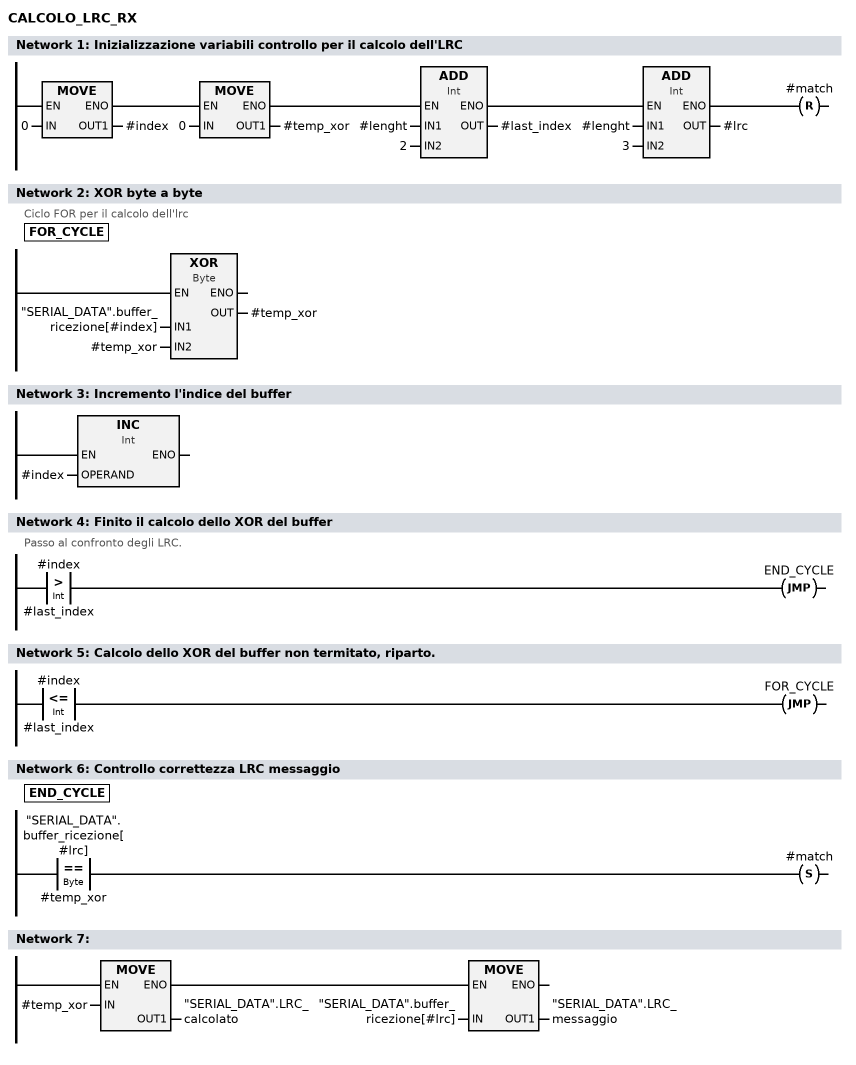
   RUNG wire#powerrail
      Move(in := 0, out1 => #index)
      Move(in := 0, out1 => #temp_xor)
      { S7_Templates := "SrcType := Int" } Add(in1 := #lenght, in2 := 2, out => #last_index)
      { S7_Templates := "SrcType := Int" } Add(in1 := #lenght, in2 := 3, out => #lrc)
      R_Coil( #match )
   END_RUNG
   // the same network as SCL:
   #index := 0;
   #temp_xor := 0;
   #last_index := #lenght + 2;
   #lrc := #lenght + 3;
   #match := FALSE;
END_REGION

REGION Network 2: XOR byte a byte
   // Ciclo FOR per il calcolo dell'lrc
   // no checked SCL form for this network; see the picture
END_REGION

REGION Network 3: Incremento l'indice del buffer
   RUNG wire#powerrail
      { S7_Templates := "DestType := Int" } Inc( #index )
   END_RUNG
   // the same network as SCL:
   #index := #index + 1;
END_REGION

REGION Network 4: Finito il calcolo dello XOR del buffer
   // Passo al confronto degli LRC.
   RUNG wire#powerrail
      { S7_Templates := "SrcType := Int" } GT_Contact(in1 := #index, in2 := #last_index)
      JumpCoil( END_CYCLE )
   END_RUNG
   // the same network as SCL:
   IF #index > #last_index THEN GOTO END_CYCLE; END_IF;
END_REGION

REGION Network 5: Calcolo dello XOR del buffer non termitato, riparto.
   RUNG wire#powerrail
      { S7_Templates := "SrcType := Int" } LE_Contact(in1 := #index, in2 := #last_index)
      JumpCoil( FOR_CYCLE )
   END_RUNG
   // the same network as SCL:
   IF #index <= #last_index THEN GOTO FOR_CYCLE; END_IF;
END_REGION

REGION Network 6: Controllo correttezza LRC messaggio
   Label( END_CYCLE )
   RUNG wire#powerrail
      { S7_Templates := "SrcType := Byte" } EQ_Contact(in1 := "SERIAL_DATA".buffer_ricezione[#lrc], in2 := #temp_xor)
      S_Coil( #match )
   END_RUNG
   // the same network as SCL:
   END_CYCLE:
   IF "SERIAL_DATA".buffer_ricezione[#lrc] = #temp_xor THEN #match := TRUE; END_IF;
END_REGION

REGION Network 7
   RUNG wire#powerrail
      Move(in := #temp_xor, out1 => "SERIAL_DATA".LRC_calcolato)
      Move(in := "SERIAL_DATA".buffer_ricezione[#lrc], out1 => "SERIAL_DATA".LRC_messaggio)
   END_RUNG
   // the same network as SCL:
   "SERIAL_DATA".LRC_calcolato := #temp_xor;
   "SERIAL_DATA".LRC_messaggio := "SERIAL_DATA".buffer_ricezione[#lrc];
END_REGION
END_FUNCTION

FUNCTION "RESET_ALLARMI" : Void   // FC7, LAD
TITLE = RESET ALLARMI
{ S7_Optimized_Access := 'FALSE' }
VERSION : 0.1
BEGIN

REGION Network 1: Azzero i contatori di fault Amplificatori
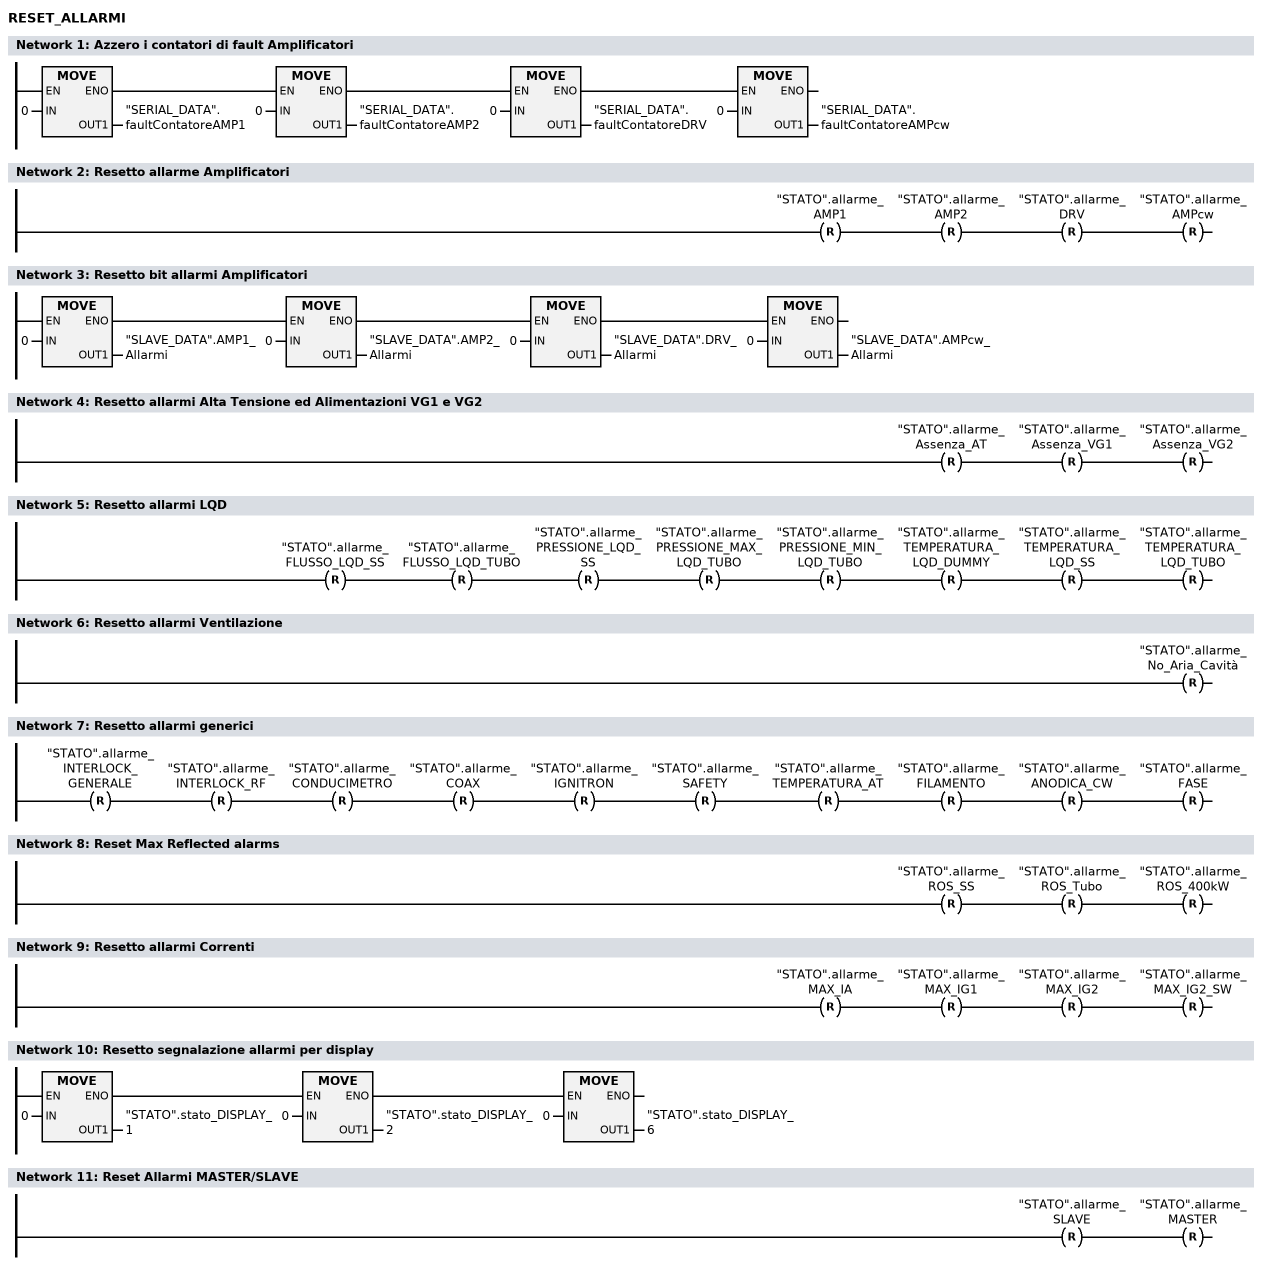
   RUNG wire#powerrail
      Move(in := 0, out1 => "SERIAL_DATA".faultContatoreAMP1)
      Move(in := 0, out1 => "SERIAL_DATA".faultContatoreAMP2)
      Move(in := 0, out1 => "SERIAL_DATA".faultContatoreDRV)
      Move(in := 0, out1 => "SERIAL_DATA".faultContatoreAMPcw)
   END_RUNG
   // the same network as SCL:
   "SERIAL_DATA".faultContatoreAMP1 := 0;
   "SERIAL_DATA".faultContatoreAMP2 := 0;
   "SERIAL_DATA".faultContatoreDRV := 0;
   "SERIAL_DATA".faultContatoreAMPcw := 0;
END_REGION

REGION Network 2: Resetto allarme Amplificatori
   RUNG wire#powerrail
      R_Coil( "STATO".allarme_AMP1 )
      R_Coil( "STATO".allarme_AMP2 )
      R_Coil( "STATO".allarme_DRV )
      R_Coil( "STATO".allarme_AMPcw )
   END_RUNG
   // the same network as SCL:
   "STATO".allarme_AMP1 := FALSE;
   "STATO".allarme_AMP2 := FALSE;
   "STATO".allarme_DRV := FALSE;
   "STATO".allarme_AMPcw := FALSE;
END_REGION

REGION Network 3: Resetto bit allarmi Amplificatori
   RUNG wire#powerrail
      Move(in := 0, out1 => "SLAVE_DATA".AMP1_Allarmi)
      Move(in := 0, out1 => "SLAVE_DATA".AMP2_Allarmi)
      Move(in := 0, out1 => "SLAVE_DATA".DRV_Allarmi)
      Move(in := 0, out1 => "SLAVE_DATA".AMPcw_Allarmi)
   END_RUNG
   // the same network as SCL:
   "SLAVE_DATA".AMP1_Allarmi := 0;
   "SLAVE_DATA".AMP2_Allarmi := 0;
   "SLAVE_DATA".DRV_Allarmi := 0;
   "SLAVE_DATA".AMPcw_Allarmi := 0;
END_REGION

REGION Network 4: Resetto allarmi Alta Tensione ed Alimentazioni VG1 e VG2
   RUNG wire#powerrail
      R_Coil( "STATO".allarme_Assenza_AT )
      R_Coil( "STATO".allarme_Assenza_VG1 )
      R_Coil( "STATO".allarme_Assenza_VG2 )
   END_RUNG
   // the same network as SCL:
   "STATO".allarme_Assenza_AT := FALSE;
   "STATO".allarme_Assenza_VG1 := FALSE;
   "STATO".allarme_Assenza_VG2 := FALSE;
END_REGION

REGION Network 5: Resetto allarmi LQD
   RUNG wire#powerrail
      R_Coil( "STATO".allarme_FLUSSO_LQD_SS )
      R_Coil( "STATO".allarme_FLUSSO_LQD_TUBO )
      R_Coil( "STATO".allarme_PRESSIONE_LQD_SS )
      R_Coil( "STATO".allarme_PRESSIONE_MAX_LQD_TUBO )
      R_Coil( "STATO".allarme_PRESSIONE_MIN_LQD_TUBO )
      R_Coil( "STATO".allarme_TEMPERATURA_LQD_DUMMY )
      R_Coil( "STATO".allarme_TEMPERATURA_LQD_SS )
      R_Coil( "STATO".allarme_TEMPERATURA_LQD_TUBO )
   END_RUNG
   // the same network as SCL:
   "STATO".allarme_FLUSSO_LQD_SS := FALSE;
   "STATO".allarme_FLUSSO_LQD_TUBO := FALSE;
   "STATO".allarme_PRESSIONE_LQD_SS := FALSE;
   "STATO".allarme_PRESSIONE_MAX_LQD_TUBO := FALSE;
   "STATO".allarme_PRESSIONE_MIN_LQD_TUBO := FALSE;
   "STATO".allarme_TEMPERATURA_LQD_DUMMY := FALSE;
   "STATO".allarme_TEMPERATURA_LQD_SS := FALSE;
   "STATO".allarme_TEMPERATURA_LQD_TUBO := FALSE;
END_REGION

REGION Network 6: Resetto allarmi Ventilazione
   RUNG wire#powerrail
      R_Coil( "STATO".allarme_No_Aria_Cavità )
   END_RUNG
   // the same network as SCL:
   "STATO".allarme_No_Aria_Cavità := FALSE;
END_REGION

REGION Network 7: Resetto allarmi generici
   RUNG wire#powerrail
      R_Coil( "STATO".allarme_INTERLOCK_GENERALE )
      R_Coil( "STATO".allarme_INTERLOCK_RF )
      R_Coil( "STATO".allarme_CONDUCIMETRO )
      R_Coil( "STATO".allarme_COAX )
      R_Coil( "STATO".allarme_IGNITRON )
      R_Coil( "STATO".allarme_SAFETY )
      R_Coil( "STATO".allarme_TEMPERATURA_AT )
      R_Coil( "STATO".allarme_FILAMENTO )
      R_Coil( "STATO".allarme_ANODICA_CW )
      R_Coil( "STATO".allarme_FASE )
   END_RUNG
   // the same network as SCL:
   "STATO".allarme_INTERLOCK_GENERALE := FALSE;
   "STATO".allarme_INTERLOCK_RF := FALSE;
   "STATO".allarme_CONDUCIMETRO := FALSE;
   "STATO".allarme_COAX := FALSE;
   "STATO".allarme_IGNITRON := FALSE;
   "STATO".allarme_SAFETY := FALSE;
   "STATO".allarme_TEMPERATURA_AT := FALSE;
   "STATO".allarme_FILAMENTO := FALSE;
   "STATO".allarme_ANODICA_CW := FALSE;
   "STATO".allarme_FASE := FALSE;
END_REGION

REGION Network 8: Reset Max Reflected alarms
   RUNG wire#powerrail
      R_Coil( "STATO".allarme_ROS_SS )
      R_Coil( "STATO".allarme_ROS_Tubo )
      R_Coil( "STATO".allarme_ROS_400kW )
   END_RUNG
   // the same network as SCL:
   "STATO".allarme_ROS_SS := FALSE;
   "STATO".allarme_ROS_Tubo := FALSE;
   "STATO".allarme_ROS_400kW := FALSE;
END_REGION

REGION Network 9: Resetto allarmi Correnti
   RUNG wire#powerrail
      R_Coil( "STATO".allarme_MAX_IA )
      R_Coil( "STATO".allarme_MAX_IG1 )
      R_Coil( "STATO".allarme_MAX_IG2 )
      R_Coil( "STATO".allarme_MAX_IG2_SW )
   END_RUNG
   // the same network as SCL:
   "STATO".allarme_MAX_IA := FALSE;
   "STATO".allarme_MAX_IG1 := FALSE;
   "STATO".allarme_MAX_IG2 := FALSE;
   "STATO".allarme_MAX_IG2_SW := FALSE;
END_REGION

REGION Network 10: Resetto segnalazione allarmi per display
   RUNG wire#powerrail
      Move(in := 0, out1 => "STATO".stato_DISPLAY_1)
      Move(in := 0, out1 => "STATO".stato_DISPLAY_2)
      Move(in := 0, out1 => "STATO".stato_DISPLAY_6)
   END_RUNG
   // the same network as SCL:
   "STATO".stato_DISPLAY_1 := 0;
   "STATO".stato_DISPLAY_2 := 0;
   "STATO".stato_DISPLAY_6 := 0;
END_REGION

REGION Network 11: Reset Allarmi MASTER/SLAVE
   RUNG wire#powerrail
      R_Coil( "STATO".allarme_SLAVE )
      R_Coil( "STATO".allarme_MASTER )
   END_RUNG
   // the same network as SCL:
   "STATO".allarme_SLAVE := FALSE;
   "STATO".allarme_MASTER := FALSE;
END_REGION
END_FUNCTION

FUNCTION "CALCOLO_LRC_TX" : Void   // FC8, LAD
TITLE = CALCOLO LRC TX
{ S7_Optimized_Access := 'FALSE' }
AUTHOR : Dario
VERSION : 0.1
// Calcolo dell'LRC per messaggi da trasmettere di tipo 49h
BEGIN

REGION Network 1: Carico indirizzo Scheda Delay
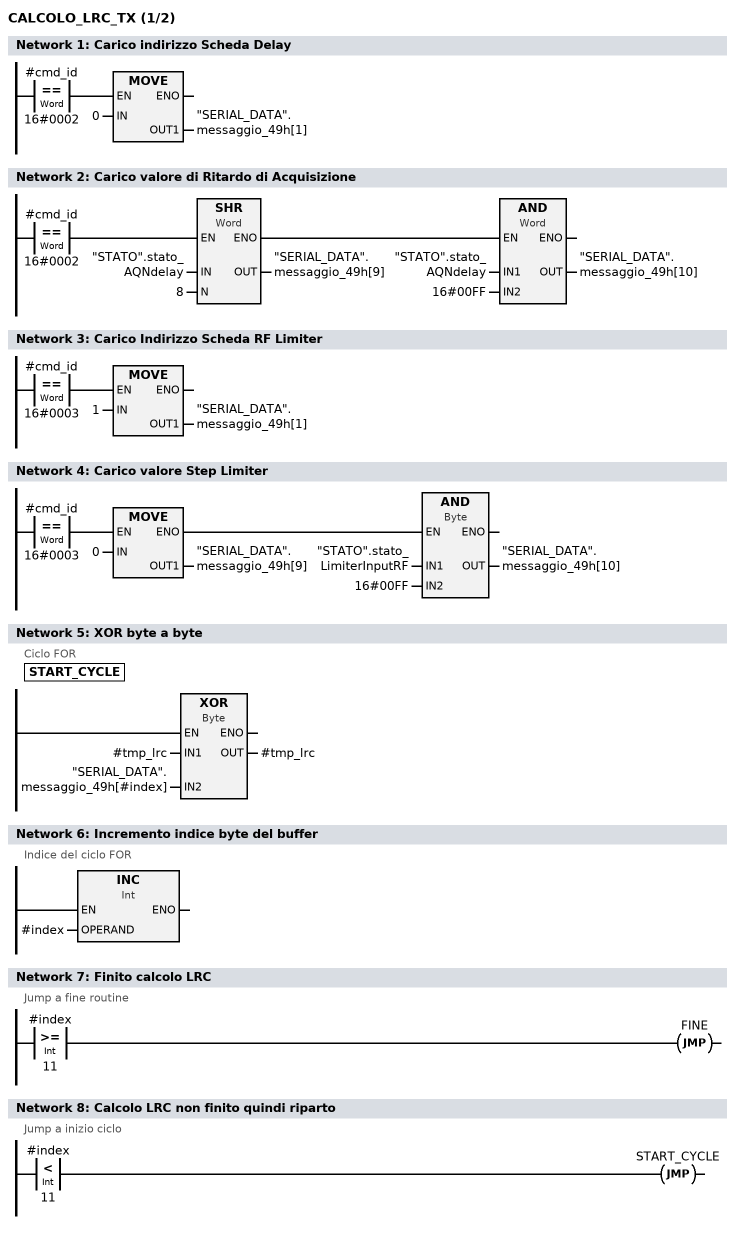
   RUNG wire#powerrail
      { S7_Templates := "SrcType := Word" } EQ_Contact(in1 := #cmd_id, in2 := 16#0002)
      Move(in := 0, out1 => "SERIAL_DATA".messaggio_49h[1])
   END_RUNG
   // the same network as SCL:
   IF #cmd_id = 16#0002 THEN "SERIAL_DATA".messaggio_49h[1] := 0; END_IF;
END_REGION

REGION Network 2: Carico valore di Ritardo di Acquisizione
   // no checked SCL form for this network; see the picture
END_REGION

REGION Network 3: Carico Indirizzo Scheda RF Limiter
   RUNG wire#powerrail
      { S7_Templates := "SrcType := Word" } EQ_Contact(in1 := #cmd_id, in2 := 16#0003)
      Move(in := 1, out1 => "SERIAL_DATA".messaggio_49h[1])
   END_RUNG
   // the same network as SCL:
   IF #cmd_id = 16#0003 THEN "SERIAL_DATA".messaggio_49h[1] := 1; END_IF;
END_REGION

REGION Network 4: Carico valore Step Limiter
   // no checked SCL form for this network; see the picture
END_REGION

REGION Network 5: XOR byte a byte
   // Ciclo FOR
   // no checked SCL form for this network; see the picture
END_REGION

REGION Network 6: Incremento indice byte del buffer
   // Indice del ciclo FOR
   RUNG wire#powerrail
      { S7_Templates := "DestType := Int" } Inc( #index )
   END_RUNG
   // the same network as SCL:
   #index := #index + 1;
END_REGION

REGION Network 7: Finito calcolo LRC
   // Jump a fine routine
   RUNG wire#powerrail
      { S7_Templates := "SrcType := Int" } GE_Contact(in1 := #index, in2 := 11)
      JumpCoil( FINE )
   END_RUNG
   // the same network as SCL:
   IF #index >= 11 THEN GOTO FINE; END_IF;
END_REGION

REGION Network 8: Calcolo LRC non finito quindi riparto
   // Jump a inizio ciclo
   RUNG wire#powerrail
      { S7_Templates := "SrcType := Int" } LT_Contact(in1 := #index, in2 := 11)
      JumpCoil( START_CYCLE )
   END_RUNG
   // the same network as SCL:
   IF #index < 11 THEN GOTO START_CYCLE; END_IF;
END_REGION

REGION Network 9: Carico l'LRC calcolato
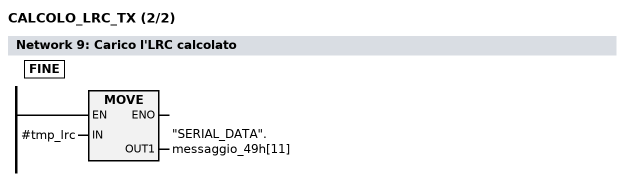
   Label( FINE )
   RUNG wire#powerrail
      Move(in := #tmp_lrc, out1 => "SERIAL_DATA".messaggio_49h[11])
   END_RUNG
   // the same network as SCL:
   FINE:
   "SERIAL_DATA".messaggio_49h[11] := #tmp_lrc;
END_REGION
END_FUNCTION

FUNCTION "SEGNALAZIONE_ALLARMI" : Void   // FC9, LAD
{ S7_Optimized_Access := 'FALSE' }
VERSION : 0.1
BEGIN

REGION Network 1: Presenza allarme flusso LQD minimo Tubo
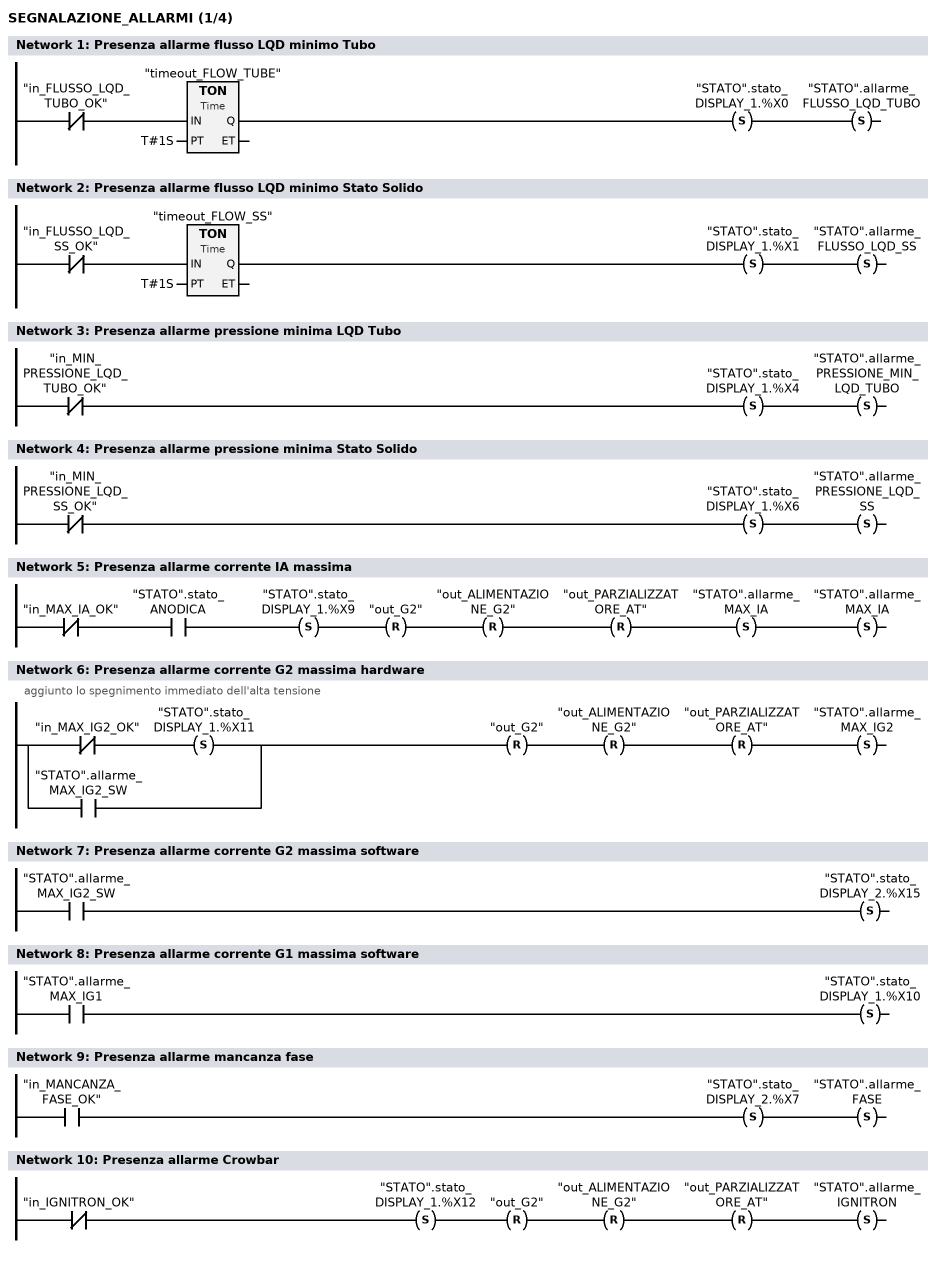
   "timeout_FLOW_TUBE".TON(IN := NOT "in_FLUSSO_LQD_TUBO_OK", PT := T#1S);
   IF "timeout_FLOW_TUBE".Q THEN
       "STATO".stato_DISPLAY_1.%X0 := TRUE;
       "STATO".allarme_FLUSSO_LQD_TUBO := TRUE;
   END_IF;
END_REGION

REGION Network 2: Presenza allarme flusso LQD minimo Stato Solido
   "timeout_FLOW_SS".TON(IN := NOT "in_FLUSSO_LQD_SS_OK", PT := T#1S);
   IF "timeout_FLOW_SS".Q THEN
       "STATO".stato_DISPLAY_1.%X1 := TRUE;
       "STATO".allarme_FLUSSO_LQD_SS := TRUE;
   END_IF;
END_REGION

REGION Network 3: Presenza allarme pressione minima LQD Tubo
   RUNG wire#powerrail
      I_Contact( "in_MIN_PRESSIONE_LQD_TUBO_OK" )
      S_Coil( "STATO".stato_DISPLAY_1.%X4 )
      S_Coil( "STATO".allarme_PRESSIONE_MIN_LQD_TUBO )
   END_RUNG
   // the same network as SCL:
   IF NOT "in_MIN_PRESSIONE_LQD_TUBO_OK" THEN
       "STATO".stato_DISPLAY_1.%X4 := TRUE;
       "STATO".allarme_PRESSIONE_MIN_LQD_TUBO := TRUE;
   END_IF;
END_REGION

REGION Network 4: Presenza allarme pressione minima Stato Solido
   RUNG wire#powerrail
      I_Contact( "in_MIN_PRESSIONE_LQD_SS_OK" )
      S_Coil( "STATO".stato_DISPLAY_1.%X6 )
      S_Coil( "STATO".allarme_PRESSIONE_LQD_SS )
   END_RUNG
   // the same network as SCL:
   IF NOT "in_MIN_PRESSIONE_LQD_SS_OK" THEN
       "STATO".stato_DISPLAY_1.%X6 := TRUE;
       "STATO".allarme_PRESSIONE_LQD_SS := TRUE;
   END_IF;
END_REGION

REGION Network 5: Presenza allarme corrente IA massima
   RUNG wire#powerrail
      I_Contact( "in_MAX_IA_OK" )
      Contact( "STATO".stato_ANODICA )
      S_Coil( "STATO".stato_DISPLAY_1.%X9 )
      R_Coil( "out_G2" )
      R_Coil( "out_ALIMENTAZIONE_G2" )
      R_Coil( "out_PARZIALIZZATORE_AT" )
      S_Coil( "STATO".allarme_MAX_IA )
      S_Coil( "STATO".allarme_MAX_IA )
   END_RUNG
   // the same network as SCL:
   IF NOT "in_MAX_IA_OK" AND "STATO".stato_ANODICA THEN
       "STATO".stato_DISPLAY_1.%X9 := TRUE;
       "out_G2" := FALSE;
       "out_ALIMENTAZIONE_G2" := FALSE;
       "out_PARZIALIZZATORE_AT" := FALSE;
       "STATO".allarme_MAX_IA := TRUE;
       "STATO".allarme_MAX_IA := TRUE;
   END_IF;
END_REGION

REGION Network 6: Presenza allarme corrente G2 massima hardware
   // aggiunto lo spegnimento immediato dell'alta tensione
   RUNG wire#powerrail
      I_Contact( "in_MAX_IG2_OK" )
      S_Coil( "STATO".stato_DISPLAY_1.%X11 )
      wire#w1
      R_Coil( "out_G2" )
      R_Coil( "out_ALIMENTAZIONE_G2" )
      R_Coil( "out_PARZIALIZZATORE_AT" )
      S_Coil( "STATO".allarme_MAX_IG2 )
   END_RUNG
   RUNG wire#powerrail
      Contact( "STATO".allarme_MAX_IG2_SW )
   END_RUNG wire#w1
   // the same network as SCL:
   IF NOT "in_MAX_IG2_OK" THEN "STATO".stato_DISPLAY_1.%X11 := TRUE; END_IF;
   IF NOT "in_MAX_IG2_OK" OR "STATO".allarme_MAX_IG2_SW THEN
       "out_G2" := FALSE;
       "out_ALIMENTAZIONE_G2" := FALSE;
       "out_PARZIALIZZATORE_AT" := FALSE;
       "STATO".allarme_MAX_IG2 := TRUE;
   END_IF;
END_REGION

REGION Network 7: Presenza allarme corrente G2 massima software
   RUNG wire#powerrail
      Contact( "STATO".allarme_MAX_IG2_SW )
      S_Coil( "STATO".stato_DISPLAY_2.%X15 )
   END_RUNG
   // the same network as SCL:
   IF "STATO".allarme_MAX_IG2_SW THEN "STATO".stato_DISPLAY_2.%X15 := TRUE; END_IF;
END_REGION

REGION Network 8: Presenza allarme corrente G1 massima software
   RUNG wire#powerrail
      Contact( "STATO".allarme_MAX_IG1 )
      S_Coil( "STATO".stato_DISPLAY_1.%X10 )
   END_RUNG
   // the same network as SCL:
   IF "STATO".allarme_MAX_IG1 THEN "STATO".stato_DISPLAY_1.%X10 := TRUE; END_IF;
END_REGION

REGION Network 9: Presenza allarme mancanza fase
   RUNG wire#powerrail
      Contact( "in_MANCANZA_FASE_OK" )
      S_Coil( "STATO".stato_DISPLAY_2.%X7 )
      S_Coil( "STATO".allarme_FASE )
   END_RUNG
   // the same network as SCL:
   IF "in_MANCANZA_FASE_OK" THEN
       "STATO".stato_DISPLAY_2.%X7 := TRUE;
       "STATO".allarme_FASE := TRUE;
   END_IF;
END_REGION

REGION Network 10: Presenza allarme Crowbar
   RUNG wire#powerrail
      I_Contact( "in_IGNITRON_OK" )
      S_Coil( "STATO".stato_DISPLAY_1.%X12 )
      R_Coil( "out_G2" )
      R_Coil( "out_ALIMENTAZIONE_G2" )
      R_Coil( "out_PARZIALIZZATORE_AT" )
      S_Coil( "STATO".allarme_IGNITRON )
   END_RUNG
   // the same network as SCL:
   IF NOT "in_IGNITRON_OK" THEN
       "STATO".stato_DISPLAY_1.%X12 := TRUE;
       "out_G2" := FALSE;
       "out_ALIMENTAZIONE_G2" := FALSE;
       "out_PARZIALIZZATORE_AT" := FALSE;
       "STATO".allarme_IGNITRON := TRUE;
   END_IF;
END_REGION

REGION Network 11: Presenza allarme Conducimetro
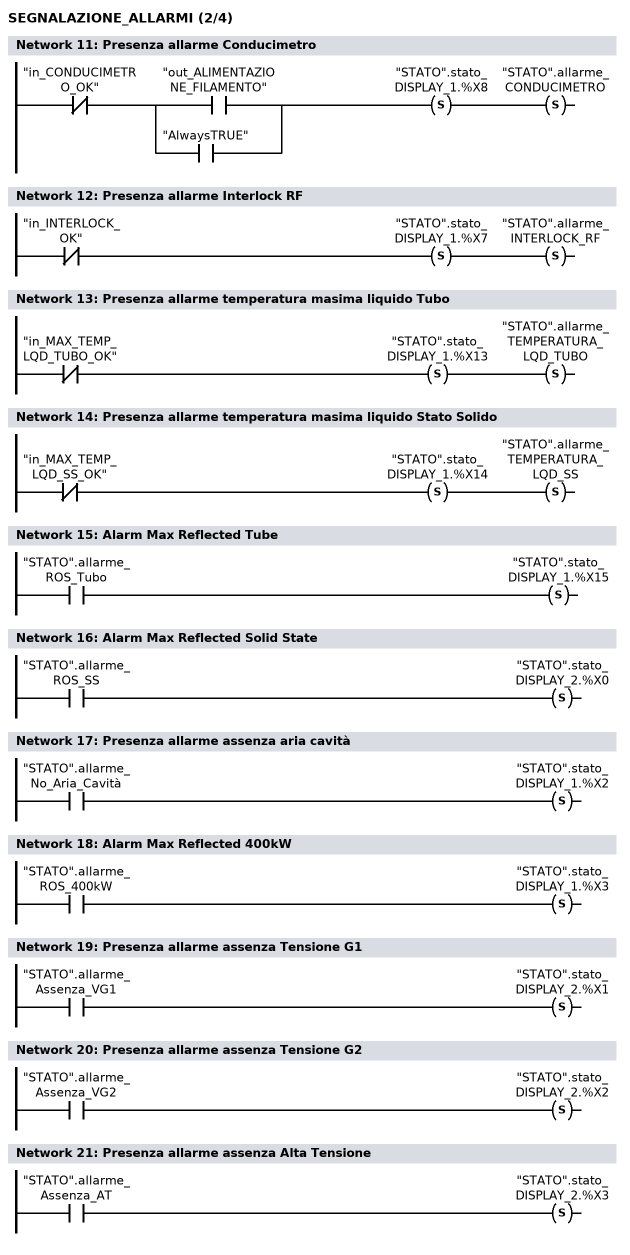
   RUNG wire#powerrail
      I_Contact( "in_CONDUCIMETRO_OK" )
      wire#w1
      Contact( "out_ALIMENTAZIONE_FILAMENTO" )
      wire#w2
      S_Coil( "STATO".stato_DISPLAY_1.%X8 )
      S_Coil( "STATO".allarme_CONDUCIMETRO )
   END_RUNG
   RUNG wire#w1
      Contact( "AlwaysTRUE" )
   END_RUNG wire#w2
   // the same network as SCL:
   IF NOT "in_CONDUCIMETRO_OK" AND ("out_ALIMENTAZIONE_FILAMENTO" OR "AlwaysTRUE") THEN
       "STATO".stato_DISPLAY_1.%X8 := TRUE;
       "STATO".allarme_CONDUCIMETRO := TRUE;
   END_IF;
END_REGION

REGION Network 12: Presenza allarme Interlock RF
   RUNG wire#powerrail
      I_Contact( "in_INTERLOCK_OK" )
      S_Coil( "STATO".stato_DISPLAY_1.%X7 )
      S_Coil( "STATO".allarme_INTERLOCK_RF )
   END_RUNG
   // the same network as SCL:
   IF NOT "in_INTERLOCK_OK" THEN
       "STATO".stato_DISPLAY_1.%X7 := TRUE;
       "STATO".allarme_INTERLOCK_RF := TRUE;
   END_IF;
END_REGION

REGION Network 13: Presenza allarme temperatura masima liquido Tubo
   RUNG wire#powerrail
      I_Contact( "in_MAX_TEMP_LQD_TUBO_OK" )
      S_Coil( "STATO".stato_DISPLAY_1.%X13 )
      S_Coil( "STATO".allarme_TEMPERATURA_LQD_TUBO )
   END_RUNG
   // the same network as SCL:
   IF NOT "in_MAX_TEMP_LQD_TUBO_OK" THEN
       "STATO".stato_DISPLAY_1.%X13 := TRUE;
       "STATO".allarme_TEMPERATURA_LQD_TUBO := TRUE;
   END_IF;
END_REGION

REGION Network 14: Presenza allarme temperatura masima liquido Stato Solido
   RUNG wire#powerrail
      I_Contact( "in_MAX_TEMP_LQD_SS_OK" )
      S_Coil( "STATO".stato_DISPLAY_1.%X14 )
      S_Coil( "STATO".allarme_TEMPERATURA_LQD_SS )
   END_RUNG
   // the same network as SCL:
   IF NOT "in_MAX_TEMP_LQD_SS_OK" THEN
       "STATO".stato_DISPLAY_1.%X14 := TRUE;
       "STATO".allarme_TEMPERATURA_LQD_SS := TRUE;
   END_IF;
END_REGION

REGION Network 15: Alarm Max Reflected Tube
   RUNG wire#powerrail
      Contact( "STATO".allarme_ROS_Tubo )
      S_Coil( "STATO".stato_DISPLAY_1.%X15 )
   END_RUNG
   // the same network as SCL:
   IF "STATO".allarme_ROS_Tubo THEN "STATO".stato_DISPLAY_1.%X15 := TRUE; END_IF;
END_REGION

REGION Network 16: Alarm Max Reflected Solid State
   RUNG wire#powerrail
      Contact( "STATO".allarme_ROS_SS )
      S_Coil( "STATO".stato_DISPLAY_2.%X0 )
   END_RUNG
   // the same network as SCL:
   IF "STATO".allarme_ROS_SS THEN "STATO".stato_DISPLAY_2.%X0 := TRUE; END_IF;
END_REGION

REGION Network 17: Presenza allarme assenza aria cavità
   RUNG wire#powerrail
      Contact( "STATO".allarme_No_Aria_Cavità )
      S_Coil( "STATO".stato_DISPLAY_1.%X2 )
   END_RUNG
   // the same network as SCL:
   IF "STATO".allarme_No_Aria_Cavità THEN "STATO".stato_DISPLAY_1.%X2 := TRUE; END_IF;
END_REGION

REGION Network 18: Alarm Max Reflected 400kW
   RUNG wire#powerrail
      Contact( "STATO".allarme_ROS_400kW )
      S_Coil( "STATO".stato_DISPLAY_1.%X3 )
   END_RUNG
   // the same network as SCL:
   IF "STATO".allarme_ROS_400kW THEN "STATO".stato_DISPLAY_1.%X3 := TRUE; END_IF;
END_REGION

REGION Network 19: Presenza allarme assenza Tensione G1
   RUNG wire#powerrail
      Contact( "STATO".allarme_Assenza_VG1 )
      S_Coil( "STATO".stato_DISPLAY_2.%X1 )
   END_RUNG
   // the same network as SCL:
   IF "STATO".allarme_Assenza_VG1 THEN "STATO".stato_DISPLAY_2.%X1 := TRUE; END_IF;
END_REGION

REGION Network 20: Presenza allarme assenza Tensione G2
   RUNG wire#powerrail
      Contact( "STATO".allarme_Assenza_VG2 )
      S_Coil( "STATO".stato_DISPLAY_2.%X2 )
   END_RUNG
   // the same network as SCL:
   IF "STATO".allarme_Assenza_VG2 THEN "STATO".stato_DISPLAY_2.%X2 := TRUE; END_IF;
END_REGION

REGION Network 21: Presenza allarme assenza Alta Tensione
   RUNG wire#powerrail
      Contact( "STATO".allarme_Assenza_AT )
      S_Coil( "STATO".stato_DISPLAY_2.%X3 )
   END_RUNG
   // the same network as SCL:
   IF "STATO".allarme_Assenza_AT THEN "STATO".stato_DISPLAY_2.%X3 := TRUE; END_IF;
END_REGION

REGION Network 22: Presenza allarme Amplificatore 1 [Impulsivo]
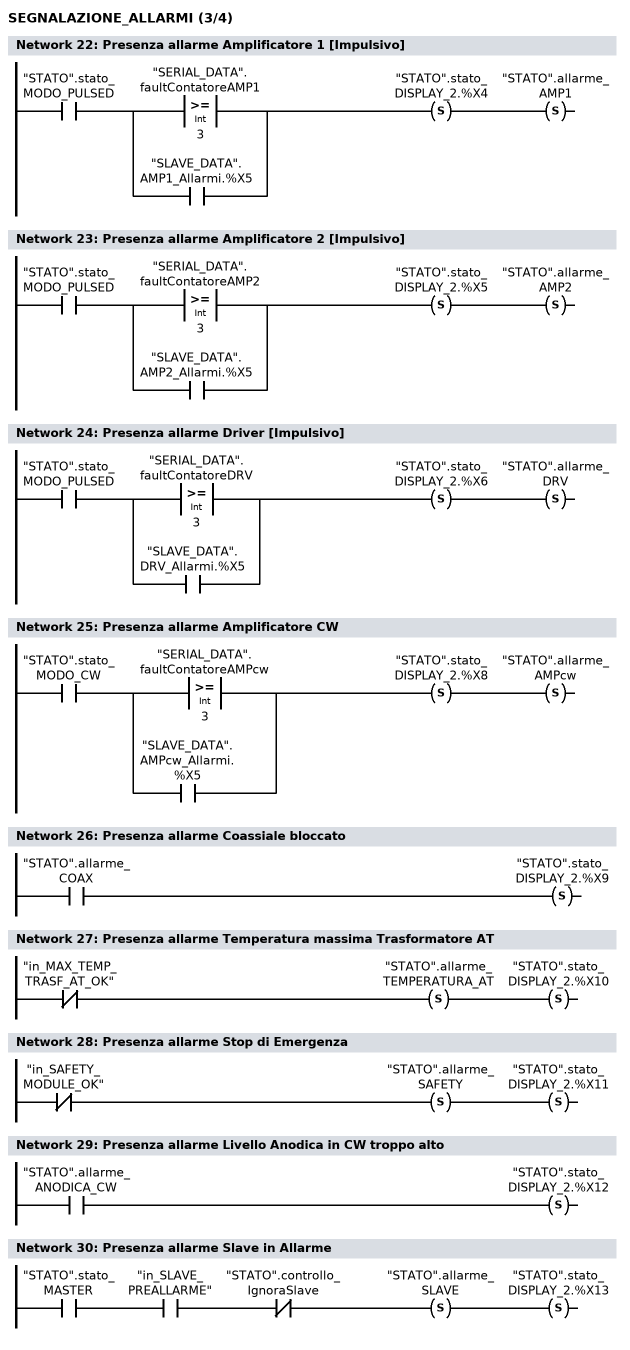
   RUNG wire#powerrail
      Contact( "STATO".stato_MODO_PULSED )
      wire#w1
      { S7_Templates := "SrcType := Int" } GE_Contact(in1 := "SERIAL_DATA".faultContatoreAMP1, in2 := 3)
      wire#w2
      S_Coil( "STATO".stato_DISPLAY_2.%X4 )
      S_Coil( "STATO".allarme_AMP1 )
   END_RUNG
   RUNG wire#w1
      Contact( "SLAVE_DATA".AMP1_Allarmi.%X5 )
   END_RUNG wire#w2
   // the same network as SCL:
   IF "STATO".stato_MODO_PULSED AND (("SERIAL_DATA".faultContatoreAMP1 >= 3) OR "SLAVE_DATA".AMP1_Allarmi.%X5) THEN
       "STATO".stato_DISPLAY_2.%X4 := TRUE;
       "STATO".allarme_AMP1 := TRUE;
   END_IF;
END_REGION

REGION Network 23: Presenza allarme Amplificatore 2 [Impulsivo]
   RUNG wire#powerrail
      Contact( "STATO".stato_MODO_PULSED )
      wire#w1
      { S7_Templates := "SrcType := Int" } GE_Contact(in1 := "SERIAL_DATA".faultContatoreAMP2, in2 := 3)
      wire#w2
      S_Coil( "STATO".stato_DISPLAY_2.%X5 )
      S_Coil( "STATO".allarme_AMP2 )
   END_RUNG
   RUNG wire#w1
      Contact( "SLAVE_DATA".AMP2_Allarmi.%X5 )
   END_RUNG wire#w2
   // the same network as SCL:
   IF "STATO".stato_MODO_PULSED AND (("SERIAL_DATA".faultContatoreAMP2 >= 3) OR "SLAVE_DATA".AMP2_Allarmi.%X5) THEN
       "STATO".stato_DISPLAY_2.%X5 := TRUE;
       "STATO".allarme_AMP2 := TRUE;
   END_IF;
END_REGION

REGION Network 24: Presenza allarme Driver [Impulsivo]
   RUNG wire#powerrail
      Contact( "STATO".stato_MODO_PULSED )
      wire#w1
      { S7_Templates := "SrcType := Int" } GE_Contact(in1 := "SERIAL_DATA".faultContatoreDRV, in2 := 3)
      wire#w2
      S_Coil( "STATO".stato_DISPLAY_2.%X6 )
      S_Coil( "STATO".allarme_DRV )
   END_RUNG
   RUNG wire#w1
      Contact( "SLAVE_DATA".DRV_Allarmi.%X5 )
   END_RUNG wire#w2
   // the same network as SCL:
   IF "STATO".stato_MODO_PULSED AND (("SERIAL_DATA".faultContatoreDRV >= 3) OR "SLAVE_DATA".DRV_Allarmi.%X5) THEN
       "STATO".stato_DISPLAY_2.%X6 := TRUE;
       "STATO".allarme_DRV := TRUE;
   END_IF;
END_REGION

REGION Network 25: Presenza allarme Amplificatore CW
   RUNG wire#powerrail
      Contact( "STATO".stato_MODO_CW )
      wire#w1
      { S7_Templates := "SrcType := Int" } GE_Contact(in1 := "SERIAL_DATA".faultContatoreAMPcw, in2 := 3)
      wire#w2
      S_Coil( "STATO".stato_DISPLAY_2.%X8 )
      S_Coil( "STATO".allarme_AMPcw )
   END_RUNG
   RUNG wire#w1
      Contact( "SLAVE_DATA".AMPcw_Allarmi.%X5 )
   END_RUNG wire#w2
   // the same network as SCL:
   IF "STATO".stato_MODO_CW AND (("SERIAL_DATA".faultContatoreAMPcw >= 3) OR "SLAVE_DATA".AMPcw_Allarmi.%X5) THEN
       "STATO".stato_DISPLAY_2.%X8 := TRUE;
       "STATO".allarme_AMPcw := TRUE;
   END_IF;
END_REGION

REGION Network 26: Presenza allarme Coassiale bloccato
   RUNG wire#powerrail
      Contact( "STATO".allarme_COAX )
      S_Coil( "STATO".stato_DISPLAY_2.%X9 )
   END_RUNG
   // the same network as SCL:
   IF "STATO".allarme_COAX THEN "STATO".stato_DISPLAY_2.%X9 := TRUE; END_IF;
END_REGION

REGION Network 27: Presenza allarme Temperatura massima Trasformatore AT
   RUNG wire#powerrail
      I_Contact( "in_MAX_TEMP_TRASF_AT_OK" )
      S_Coil( "STATO".allarme_TEMPERATURA_AT )
      S_Coil( "STATO".stato_DISPLAY_2.%X10 )
   END_RUNG
   // the same network as SCL:
   IF NOT "in_MAX_TEMP_TRASF_AT_OK" THEN
       "STATO".allarme_TEMPERATURA_AT := TRUE;
       "STATO".stato_DISPLAY_2.%X10 := TRUE;
   END_IF;
END_REGION

REGION Network 28: Presenza allarme Stop di Emergenza
   RUNG wire#powerrail
      I_Contact( "in_SAFETY_MODULE_OK" )
      S_Coil( "STATO".allarme_SAFETY )
      S_Coil( "STATO".stato_DISPLAY_2.%X11 )
   END_RUNG
   // the same network as SCL:
   IF NOT "in_SAFETY_MODULE_OK" THEN
       "STATO".allarme_SAFETY := TRUE;
       "STATO".stato_DISPLAY_2.%X11 := TRUE;
   END_IF;
END_REGION

REGION Network 29: Presenza allarme Livello Anodica in CW troppo alto
   RUNG wire#powerrail
      Contact( "STATO".allarme_ANODICA_CW )
      S_Coil( "STATO".stato_DISPLAY_2.%X12 )
   END_RUNG
   // the same network as SCL:
   IF "STATO".allarme_ANODICA_CW THEN "STATO".stato_DISPLAY_2.%X12 := TRUE; END_IF;
END_REGION

REGION Network 30: Presenza allarme Slave in Allarme
   RUNG wire#powerrail
      Contact( "STATO".stato_MASTER )
      Contact( "in_SLAVE_PREALLARME" )
      I_Contact( "STATO".controllo_IgnoraSlave )
      S_Coil( "STATO".allarme_SLAVE )
      S_Coil( "STATO".stato_DISPLAY_2.%X13 )
   END_RUNG
   // the same network as SCL:
   IF "STATO".stato_MASTER AND "in_SLAVE_PREALLARME" AND NOT "STATO".controllo_IgnoraSlave THEN
       "STATO".allarme_SLAVE := TRUE;
       "STATO".stato_DISPLAY_2.%X13 := TRUE;
   END_IF;
END_REGION

REGION Network 31: Presenza allarme Slave in Blocco
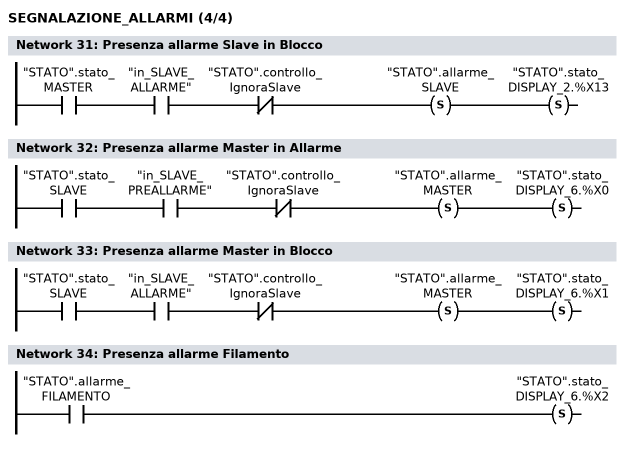
   RUNG wire#powerrail
      Contact( "STATO".stato_MASTER )
      Contact( "in_SLAVE_ALLARME" )
      I_Contact( "STATO".controllo_IgnoraSlave )
      S_Coil( "STATO".allarme_SLAVE )
      S_Coil( "STATO".stato_DISPLAY_2.%X13 )
   END_RUNG
   // the same network as SCL:
   IF "STATO".stato_MASTER AND "in_SLAVE_ALLARME" AND NOT "STATO".controllo_IgnoraSlave THEN
       "STATO".allarme_SLAVE := TRUE;
       "STATO".stato_DISPLAY_2.%X13 := TRUE;
   END_IF;
END_REGION

REGION Network 32: Presenza allarme Master in Allarme
   RUNG wire#powerrail
      Contact( "STATO".stato_SLAVE )
      Contact( "in_SLAVE_PREALLARME" )
      I_Contact( "STATO".controllo_IgnoraSlave )
      S_Coil( "STATO".allarme_MASTER )
      S_Coil( "STATO".stato_DISPLAY_6.%X0 )
   END_RUNG
   // the same network as SCL:
   IF "STATO".stato_SLAVE AND "in_SLAVE_PREALLARME" AND NOT "STATO".controllo_IgnoraSlave THEN
       "STATO".allarme_MASTER := TRUE;
       "STATO".stato_DISPLAY_6.%X0 := TRUE;
   END_IF;
END_REGION

REGION Network 33: Presenza allarme Master in Blocco
   RUNG wire#powerrail
      Contact( "STATO".stato_SLAVE )
      Contact( "in_SLAVE_ALLARME" )
      I_Contact( "STATO".controllo_IgnoraSlave )
      S_Coil( "STATO".allarme_MASTER )
      S_Coil( "STATO".stato_DISPLAY_6.%X1 )
   END_RUNG
   // the same network as SCL:
   IF "STATO".stato_SLAVE AND "in_SLAVE_ALLARME" AND NOT "STATO".controllo_IgnoraSlave THEN
       "STATO".allarme_MASTER := TRUE;
       "STATO".stato_DISPLAY_6.%X1 := TRUE;
   END_IF;
END_REGION

REGION Network 34: Presenza allarme Filamento
   RUNG wire#powerrail
      Contact( "STATO".allarme_FILAMENTO )
      S_Coil( "STATO".stato_DISPLAY_6.%X2 )
   END_RUNG
   // the same network as SCL:
   IF "STATO".allarme_FILAMENTO THEN "STATO".stato_DISPLAY_6.%X2 := TRUE; END_IF;
END_REGION
END_FUNCTION

FUNCTION "AGGIORNO_EVENTI" : Void   // FC10, LAD
{ S7_Optimized_Access := 'FALSE' }
VERSION : 0.1
BEGIN

REGION Network 1: Aggiorno stato Impulsivo
   // stato_DISPLY_3.x0 = 1 è impulsivo
